
         CALL  BLKMOV
         ( SRCBLK  := "DB919_ShotResultMach".ShotResult_Ma[1],
           RET_VAL := #"Return",
           DSTBLK  := "DB919_ShotResultMach".ShotResult_Ma[0]
         );

   // Verbrauchszähler erhöhen
         CALL  "PartCounter";
         SET;
         =     "DB_Zaehler_Anzeige".Read;

         A     "DB123_MH_IO_Signals".MH[1].IN.MH_Auto_Mode;
         S     "M_NewShotDataToMC";  // For traceability
   //-
         A     "BufferShotResultM1";
         S     "DB919_ShotResultMach".ShotResult_Ma[0].General.SendData;

   m1:   NOP   0;


         AN    "DB919_ShotResultMach".ShotResult_Ma[0].General.SendData;
         R     "BufferShotResultM1";
END_REGION

REGION Network 4: PartCounter
         A     "DB_Zaehler_Anzeige".Schichtwechsel;
         JCN   Migra_CC_0;
         CALL  "PartCounterCopy";
   Migra_CC_0:SET;
         CALL  "PartCounterView";
END_REGION
END_FUNCTION_BLOCK

FUNCTION_BLOCK "FB930_FoamingData"   // FB930, STL
TITLE = Tool-Allocation -> Read tooldata and recipedata
{ S7_Optimized_Access := 'FALSE' }
AUTHOR : KT242
VERSION : 0.1
BEGIN

REGION Network 2
         CALL  "GetToolShotValues", "GetToolShotValues_DB"
         ( IN_ResetFaults    := "DB009_Faults".Faults_Reset_FKT_M1,
           IN_MachineNo      := 1,
           IN_EnableTool     := 1,
           IO_Faults         := "DB829_Error_Machine".PouringCycle[1],
           IO_FaultLevel_1   := "DB009_Faults".Faults_FKT_Grp_1_M1,
           IO_FaultLevel_2   := "DB009_Faults".Faults_FKT_Grp_2_M1,
           IO_FaultLevel_3   := "DB009_Faults".Faults_FKT_Grp_3_M1,
           IO_NewFault       := "DB009_Faults".Faultschanging_M1,
           IO_FaultAtStation := ,
           IO_PartShotNoNew  :=
         );
   //-----
END_REGION
END_FUNCTION_BLOCK

FUNCTION_BLOCK "FB1025_Service"   // FB1025, STL
{ S7_Optimized_Access := 'FALSE' }
VERSION : 0.1
   VAR_TEMP
      Inputbyte : Byte;
      Error : Word;
   END_VAR
BEGIN

REGION Network 1: Read input byte
         L     "DB1025_Service".Set.Inputbyte;
         SLW   3;
         LAR1;

         L     IB [ AR1 , P#0.0 ];
         T     "DB1025_Service".State.Inputbyte;
END_REGION

REGION Network 2: Read output byte
         L     "DB1025_Service".Set.Outputbyte;
         SLW   3;
         LAR1;

         L     QB [ AR1 , P#0.0 ];
         T     "DB1025_Service".State.Outputbyte;
END_REGION
END_FUNCTION_BLOCK

FUNCTION_BLOCK "FB1900_IF_Robots"   // FB1900, STL
TITLE = Interface Robots
{ S7_Optimized_Access := 'FALSE' }
VERSION : 0.1
   VAR_TEMP
      Auto : Bool;
      Start_cyle : Bool;
      Auto_Stop_quitt : Bool;
      Shotrelease : Bool;
      Freigabe_Eintrag_von_PUC : Bool;
      Start_Zyklus_Roboter : Bool;
      Temp_CleaningRequest : Bool;
      Temp_EnableDoorOpen : Bool;
      Automatik_Stop_ist_Quitt : Bool;
      Temp_StartCycle : Bool;
      Temp_EnableMCatPos1 : Bool;
      Temp_TestShoActiv : Bool;
      Temp_ArPos1or2 : Bool;
      Temp_FlagStartButton : Bool;
   END_VAR
BEGIN

REGION Network 1: Saftey Door 1
         ON    "DB619_State_MPart".Operationmode[1].Auto;
         ON    "DB123_MH_IO_Signals".MH[1].IN.MH_Auto_Mode;
         =     #Temp_EnableDoorOpen;
   //-----
         CALL  "FC1033_SafetyDevice"
         ( IN_With_Safety_door := true,
           IN_EnableDoorOpen   := #Temp_EnableDoorOpen,
           IN_SelectDoorOpen   := "S_SelectDoor_Robot_01",
           IN_AS_Door          := "AS_Door_Robot_01",
           IN_QuitDoorOpen     := "S_QuittDoor_Robot_01",
           IN_OMLampTest       := "DB619_State_MPart".Operationmode[1].Lamptest,
           IN_Delay_QuitDoor   := "TM_Delay_Safetydoor_1",
           OUT_V_DoorOpen      := "V_OpenDoor_Robot_01",
           OUT_H_DoorOpen      := "H_ReleaseDoor_Robot_01",
           StatusSafetyDevice  := "DB1031_AddStatus".SaftyDevice[1]
         );
   //-----
END_REGION

REGION Network 2: Saftey Door 2
         ON    "DB619_State_MPart".Operationmode[1].Auto;
         ON    "DB123_MH_IO_Signals".MH[1].IN.MH_Auto_Mode;
         =     #Temp_EnableDoorOpen;
   //-----
         CALL  "FC1033_SafetyDevice"
         ( IN_With_Safety_door := true,
           IN_EnableDoorOpen   := #Temp_EnableDoorOpen,
           IN_SelectDoorOpen   := "S_SelectDoor_TestShot_01",
           IN_AS_Door          := "AS_Door_TestShot_01",
           IN_QuitDoorOpen     := "S_QuittDoor_TestShot_01",
           IN_OMLampTest       := "DB619_State_MPart".Operationmode[1].Lamptest,
           IN_Delay_QuitDoor   := "TM_Delay_Safetydoor_2",
           OUT_V_DoorOpen      := "V_OpenDoor_TestShot_01",
           OUT_H_DoorOpen      := "H_ReleaseDoor_TestShot_01",
           StatusSafetyDevice  := "DB1031_AddStatus".SaftyDevice[2]
         );
   //-----
END_REGION

REGION Network 3: General release
         A     "AS";
         A     "DB619_State_MPart".Operationmode[1].Controllvoltage;
         A     "DB619_State_MPart".Operationmode[1].Auto;
         A     "DB123_MH_IO_Signals".MH[1].IN.MH_Auto_Mode;
         =     #Auto;
   //
         A     "AS";
         A     "DB619_State_MPart".Operationmode[1].Controllvoltage;
         =     #Auto_Stop_quitt;
   //
         AN    "AS";
         A     "DB619_State_MPart".Operationmode[1].Controllvoltage;
         A     "DB619_State_MPart".Operationmode[1].Auto;
         A     "DB123_MH_IO_Signals".MH[1].IN.MH_Auto_Mode;
         =     "DB1010_TT_Fault".AS.AS_Activ;
   //
         A     "DB619_State_MPart".Cycle[1].Release;
         =     #Shotrelease;

   // Cleaning after shot
   //-----
         A     "DB614_MH_State".MH_CleaningPiston[1].CleanAfterShotSelected;
         S     "DB1900_IF_Robots".State_Robots[1].CleaningMHRequested;
   //-
         A(;
         L     "DB1900_IF_Robots".Switch_Robots[1].StateCleaning;
         L     1;
         ==I;
         );
         R     "DB1900_IF_Robots".State_Robots[1].CleaningMHRequested;
   //-
         A     "DB1900_IF_Robots".State_Robots[1].CleaningMHRequested;
         =     #Temp_CleaningRequest;
   //-----
         CALL  "FC5901_generalFunction"
         ( StartCycle     := #Temp_StartCycle,
           EnableMCatPos1 := #Temp_EnableMCatPos1,
           TestShotActiv  := "DB1900_IF_Robots".State_Robots[1].TestShotRunning,
           AtPos1or2      := "DB1900_IF_Robots".State_Robots[1].AtPos1or2  // #Temp_ArPos1or2
         );
   //
         A     "DB1900_IF_Robots".State_Robots[1].AtPos1or2;
         =     #Temp_ArPos1or2;
END_REGION

REGION Network 4: ProgNo send to robot KUKA
         L     "DB110_Interf_Program_M1".Signals_ExPlant[1].PrgNo;
         T     "DB1900_IF_Robots".State_Kuka[1].A_SPS_PGNO;
END_REGION

REGION Network 5: Robot interface KUKA
         AN    "DB1901_Config_Robots".Config_Robots[1].Type_Kuka;
         JC    Rob_ABB;
   //------
   // Start Cycle
   //
         A     "DB110_Interf_Program_M1".Signals_ExPlant[1].cycle_run;
         FP    "FHM_PU_cycle_running";
         S     "Flag_PU_cycle_running";

         ON    "DB619_State_MPart".Cycle[1].running;
         O     "DB1900_IF_Robots".State_Kuka[1].Input_From_Robot.E_KRC_MH_OPEN;
         O     "DB1900_IF_Robots".State_Kuka[1].Input_From_Robot.E_KRC_FLT_WaitTime;
         R     "Flag_PU_cycle_running";

         A(;
         L     "DB1900_IF_Robots".State_Kuka[1].A_SPS_PGNO;
         L     0;
         >I;
         );
         A     "DB1900_IF_Robots".State_Kuka[1].Input_From_Robot.E_KRC_PGNO_REQ;
         A     "DB1900_IF_Robots".State_Kuka[1].Input_From_Robot.E_KRC_PERI_RDY;
         A     "DB1900_IF_Robots".State_Kuka[1].Input_From_Robot.E_KRC_ALARM_STOP;
         A     "DB1900_IF_Robots".State_Kuka[1].Input_From_Robot.E_KRC_USER_SAF;
         A     "DB1900_IF_Robots".State_Kuka[1].Input_From_Robot.E_KRC_AUT_EXTERN;
         A     "DB1900_IF_Robots".State_Kuka[1].Input_From_Robot.E_KRC_IN_HOME;
         A     "Flag_PU_cycle_running";
         =     #Start_cyle;


         CALL  "FC1900_IF_Kuka_KRC4"
         ( IN_PW_INOUT           := 700,
           IN_Acknowledge_Fault  := "DB009_Faults".Faults_Reset_FKT_M1,
           IN_Auto_Stop_quitt    := #Auto_Stop_quitt,
           IN_Motorprotection    := "F_Robot_01",
           IN_MH_Automatic       := #Auto,
           IN_OM_service         := "DB614_MH_State".MH_Status[1].Switch_Service_ON_OFF,
           IN_Cycle_running      := "DB619_State_MPart".Cycle[1].running,
           IN_Start_cycle        := #Start_cyle,
           IN_Release_move_MC    := TRUE,
           IN_Shotrelease        := #Shotrelease,  //"DB619_State_MPart".Cycle[1].Shotrelease
           IN_Shotend            := "DB110_Interf_Program_M1".Bits.PulseShotEnd,
           IN_FLT_Group_1        := "DB009_Faults".Fault_State_Grp_1_M1,
           IN_PGNO_MainPos       := 250,
           IN_PGNO_Cleaning      := 251,
           IN_Timer_Auto_on      := "TM_1_Robot_1",
           IN_Timer_Fault_quitt  := "TM_2_Robot_1",
           IN_Timer_Auto_On_Off  := "TM_3_Robot_1",
           IN_Timer_Delay_Start  := "TM_4_Robot_1",
           IN_Timer_PGNO_Valid   := "TM_5_Robot_1",
           IN_Timer_Imp_ExtStart := "TM_6_Robot_1",
           AB_KUKA_PGNO          := "DB1900_IF_Robots".State_Kuka[1].Output_To_Robot.A_SPS_PGNO,
           IO_Button_MainPos     := "DB1900_IF_Robots".Switch_Robots[1].SwitchMaintPosON_OFF,
           IO_Button_Cleaning    := "DB1900_IF_Robots".Switch_Robots[1].SwitchCleaningON_OFF,
           IO_State_MainPos      := "DB1900_IF_Robots".Switch_Robots[1].StateMaintPos,
           IO_State_Cleaning     := "DB1900_IF_Robots".Switch_Robots[1].StateCleaning,
           IO_Status             := "DB1900_IF_Robots".State_Kuka[1],
           IO_NewFault           := "DB009_Faults".Faultschanging_M1,
           IO_FaultLevel_3       := "DB009_Faults".Faults_FKT_Grp_3_M1
         );

   Rob_ABB:NOP   0;
END_REGION

REGION Network 6: Robot interface ABB
         AN    "DB1901_Config_Robots".Config_Robots[1].Type_ABB;
         JC    Rob_Fanuc;
   //-----
         A     "DB1900_IF_Robots".State_ABB[1].doShotDigOut_open_MH;
         A     "DB614_MH_State".MH_Status[1].OpenMHEnableExtern;
         =     "DB614_MH_State".MH_Status[1].OpenMHEnableExtern;
   //-----
   //-
         A     "DB619_State_MPart".Operationmode[1].Controllvoltage;
         =     "DB1900_IF_Robots".State_Robots[1].EmergencyStopReady;
   //-
         A     #Auto_Stop_quitt;
         =     "DB1900_IF_Robots".State_Robots[1].AutomatcStopReady;
   //-
         A     "DB619_State_MPart".Operationmode[1].Auto;
         =     "DB1900_IF_Robots".State_Robots[1].MaschineAuto;
   //-
         A     "DB123_MH_IO_Signals".MH[1].IN.MH_Auto_Mode;
         =     "DB1900_IF_Robots".State_Robots[1].MixingheadAuto;
   //-
   // Status auch in FC irgendwann!

         A     "DB1900_IF_Robots".State_ABB[1].Output.doIRBInHome;
         =     "DB1900_IF_Robots".State_Robots[1].Rob_in_Home;

         A     "DB1900_IF_Robots".State_ABB[1].Output.doIRBinAuto;
         =     "DB1900_IF_Robots".State_Robots[1].Rob_in_Automatic;

         A     "DB1900_IF_Robots".State_ABB[1].Output.doCycleStarted;
         =     "DB1900_IF_Robots".State_Robots[1].Rob_in_Cycle;

         A     "DB1900_IF_Robots".State_ABB[1].Output.doIRBinAuto;
         A     "DB1900_IF_Robots".State_ABB[1].Output.doIRBInHome;
         A     "DB1900_IF_Robots".State_ABB[1].Output.doCycleEnd;
         A(;
         L     "DB1900_IF_Robots".State_ABB[1].Stepnumber;
         L     0;
         ==I;
         );
         =     "DB1900_IF_Robots".State_Robots[1].ReadyForStartCycle;

         L     "DB1900_IF_Robots".State_ABB[1].Stepnumber;
         T     "DB1900_IF_Robots".State_Robots[1].StepNo;

         L     "DB1900_IF_Robots".State_ABB[1].Output.GOError;
         T     "DB1900_IF_Robots".State_Robots[1].FaultNo;
   ///----------
   // Not- Aus und Automatik Stop wurden quittiert:
   ///----------
         AN    "DB1900_IF_Robots".State_ABB[1].Output.doSysError;
         AN    "DB1900_IF_Robots".State_ABB[1].Output.doEmStop_Akt;
         AN    "DB1900_IF_Robots".State_ABB[1].Input.diQuickStop;
         AN    "DB1900_IF_Robots".State_ABB[1].Output.doSafeZoneActiv;
         A     #Auto_Stop_quitt;
         A     "DB123_MH_IO_Signals".MH[1].IN.MH_Auto_Mode;
         =     #Automatik_Stop_ist_Quitt;
   ///----------
   // Datenaustausch mit dem Roboter starten:
   ///----------
         A     #Temp_StartCycle;
         A     #Automatik_Stop_ist_Quitt;
         A     "DB1900_IF_Robots".State_ABB[1].Output.doIRBInHome;
         A     "DB1900_IF_Robots".State_ABB[1].Output.doIRBinAuto;
         A     "DB1900_IF_Robots".State_ABB[1].Output.doCycleOn;
         AN    "DB1900_IF_Robots".State_ABB[1].Output.doSysError;
         AN    "DB619_State_MPart".Operationmode[1].Test;
         =     #Start_Zyklus_Roboter;
   ///----------
   // Bewegungefreigabe zum Verfahren in die Formträger
   ///----------
         A     #Temp_EnableMCatPos1;
         A     "DB123_MH_IO_Signals".MH[1].IN.MH_Auto_Mode;
         AN    "DB619_State_MPart".Operationmode[1].Test;
         A     "DB619_State_MPart".Cycle[1].Shotrelease;
   //U     "DB005_RS<->Extern".MC_Interface[1].FromMC.EnableFoaming
         =     "DB1900_IF_Robots".State_ABB[1].Input.diStartMoveMC;
   //--------------------------------------------------------------------
   // Das öffnen des Mischkopfes kann von dem Roboter angesteuert werden:
   // Roboter wartet in Vorposition bis das Signal kommt.
         A     #Temp_EnableMCatPos1;
         A     "DB619_State_MPart".Cycle[1].Shotrelease;
         =     #Freigabe_Eintrag_von_PUC;
   ///----------
   // Roboter zur Maintenanceposition und zurück zur Homeposition
   ///----------
         A     "DB1900_IF_Robots".Switch_Robots[1].SwitchMaintPosON_OFF;
         A     "DB123_MH_IO_Signals".MH[1].IN.MH_Auto_Mode;
         AN    #Temp_ArPos1or2;
         A     #Automatik_Stop_ist_Quitt;  // NotHalt ???
         A     "DB1900_IF_Robots".State_ABB[1].Output.doIRBInHome;
         A     "DB1900_IF_Robots".State_ABB[1].Output.doCycleEnd;
         AN    "DB1900_IF_Robots".State_ABB[1].Output.doCycleStarted;
         S     "DB1900_IF_Robots".State_ABB[1].Input.diHomeToMaintP;
   ///----------
         O     "DB1900_IF_Robots".State_ABB[1].Output.doIRBInMaintP;
         ON    "DB1900_IF_Robots".State_ABB[1].Output.doIRBinAuto;
         ON    "DB1900_IF_Robots".State_ABB[1].Output.doCycleOn;
         R     "DB1900_IF_Robots".State_ABB[1].Input.diHomeToMaintP;
   ///----------
         AN    "DB1900_IF_Robots".Switch_Robots[1].SwitchMaintPosON_OFF;
         A     "DB123_MH_IO_Signals".MH[1].IN.MH_Auto_Mode;
         A     #Automatik_Stop_ist_Quitt;
         A     "DB1900_IF_Robots".State_ABB[1].Output.doIRBInMaintP;
         A     "DB1900_IF_Robots".State_ABB[1].Output.doCycleEnd;
         AN    "DB1900_IF_Robots".State_ABB[1].Output.doCycleStarted;
         S     "DB1900_IF_Robots".State_ABB[1].Input.diMaintToHomeP;
   ///----------
         O     "DB1900_IF_Robots".State_ABB[1].Output.doIRBInHome;
         ON    "DB1900_IF_Robots".State_ABB[1].Output.doIRBinAuto;
         ON    "DB1900_IF_Robots".State_ABB[1].Output.doCycleOn;
         R     "DB1900_IF_Robots".State_ABB[1].Input.diMaintToHomeP;
   //-----
         L     1;  // Green
         A     "DB1900_IF_Robots".State_ABB[1].Output.doIRBInMaintP;
         JC    StateMaintPos;
         L     3;  // Yellow
         O     "DB1900_IF_Robots".Switch_Robots[1].SwitchMaintPosON_OFF;
         O     "DB1900_IF_Robots".State_ABB[1].Input.diMaintToHomeP;
         JC    StateMaintPos;
         L     0;  // OFF
   StateMaintPos:NOP   0;
         T     "DB1900_IF_Robots".Switch_Robots[1].StateMaintPos;

   ///----------
   // Roboter zur 2. Maintenanceposition und zurück zur Homeposition
   ///----------
         A     "DB1900_IF_Robots".Switch_Robots[1].SwitchMaintPos_2ON_OFF;
         A     "DB123_MH_IO_Signals".MH[1].IN.MH_Auto_Mode;
         AN    #Temp_ArPos1or2;
         A     #Automatik_Stop_ist_Quitt;  // NotHalt ???
         A     "DB1900_IF_Robots".State_ABB[1].Output.doIRBInHome;
         A     "DB1900_IF_Robots".State_ABB[1].Output.doCycleEnd;
         AN    "DB1900_IF_Robots".State_ABB[1].Output.doCycleStarted;
         S     "DB1900_IF_Robots".State_ABB[1].Input.diHomeToMaint2;
   ///----------
         O     "DB1900_IF_Robots".State_ABB[1].Output.doIRBInMaintP2;
         ON    "DB1900_IF_Robots".State_ABB[1].Output.doIRBinAuto;
         ON    "DB1900_IF_Robots".State_ABB[1].Output.doCycleOn;
         R     "DB1900_IF_Robots".State_ABB[1].Input.diHomeToMaint2;
   ///----------
         AN    "DB1900_IF_Robots".Switch_Robots[1].SwitchMaintPos_2ON_OFF;
         A     "DB123_MH_IO_Signals".MH[1].IN.MH_Auto_Mode;
         A     #Automatik_Stop_ist_Quitt;
         A     "DB1900_IF_Robots".State_ABB[1].Output.doIRBInMaintP2;
         A     "DB1900_IF_Robots".State_ABB[1].Output.doCycleEnd;
         AN    "DB1900_IF_Robots".State_ABB[1].Output.doCycleStarted;
         S     "DB1900_IF_Robots".State_ABB[1].Input.diMaintToHome2;
   ///----------
         O     "DB1900_IF_Robots".State_ABB[1].Output.doIRBInHome;
         ON    "DB1900_IF_Robots".State_ABB[1].Output.doIRBinAuto;
         ON    "DB1900_IF_Robots".State_ABB[1].Output.doCycleOn;
         R     "DB1900_IF_Robots".State_ABB[1].Input.diMaintToHome2;
   //-----

         L     1;  // Green
         A     "DB1900_IF_Robots".State_ABB[1].Output.doIRBInMaintP2;
         JC    StateMaintPos2;
         L     3;  // Yellow
         O     "DB1900_IF_Robots".Switch_Robots[1].SwitchMaintPos_2ON_OFF;
         O     "DB1900_IF_Robots".State_ABB[1].Input.diMaintToHome2;
         JC    StateMaintPos2;
         L     0;  // OFF
   StateMaintPos2:NOP   0;
         T     "DB1900_IF_Robots".Switch_Robots[1].StateMaintPos_2;

   //-----
   // Robot to mixinghead cleaning
   //-----
         A(;
         A     "DB1900_IF_Robots".Switch_Robots[1].SwitchBrushON_OFF;
         AN    #Temp_ArPos1or2;
         A     "DB1900_IF_Robots".State_ABB[1].Output.doIRBInHome;
         A     "DB1900_IF_Robots".State_ABB[1].Output.doCycleEnd;
         AN    "DB1900_IF_Robots".State_ABB[1].Output.doCycleStarted;
         O;
         A     "DB619_State_MPart".Cycle[1].ShotRuns;
         A     "DB614_MH_State".MH_CleaningPiston[1].CleanAfterShotSelected;
         );
         A     #Automatik_Stop_ist_Quitt;
         S     "DB1900_IF_Robots".State_ABB[1].Input.diStartBrushMH;
         S     "DB1900_IF_Robots".State_ABB[1].CleaningSelected;
   //-----
         O     "DB1900_IF_Robots".State_ABB[1].Output.doCleanBrushOn;
         ON    "DB1900_IF_Robots".State_ABB[1].Output.doIRBinAuto;
         ON    "DB1900_IF_Robots".State_ABB[1].Output.doCycleOn;
         R     "DB1900_IF_Robots".State_ABB[1].Input.diStartBrushMH;
   //-----
         A     "DB1900_IF_Robots".State_ABB[1].Output.doCleanBrushOn;
         FN    "DB1900_IF_Robots".State_ABB[1].FHM_CleaningActiv;
         =     "DB1900_IF_Robots".State_ABB[1].CleaningActiv;
   //-----
         A     "DB1900_IF_Robots".State_ABB[1].CleaningActiv;
         R     "DB1900_IF_Robots".State_ABB[1].CleaningSelected;
         R     "DB1900_IF_Robots".Switch_Robots[1].SwitchBrushON_OFF;
   //-----
   // Ansteuerung des Reinigungskolben vom Roboter aus
         A     "DB1900_IF_Robots".State_ABB[1].Output.doCleanBrushOn;
         =     "DB1900_IF_Robots".State_Robots[1].CleaningMHOn;
   //-----
         L     1;  // Green
         A     "DB1900_IF_Robots".State_ABB[1].Output.doCleanBrushOn;
         JC    StateCleaningMH;
         L     3;  // Yellow
         O     "DB1900_IF_Robots".Switch_Robots[1].SwitchBrushON_OFF;
         O     "DB1900_IF_Robots".State_ABB[1].CleaningSelected;
         JC    StateCleaningMH;
         L     0;  // OFF
   StateCleaningMH:NOP   0;
         T     "DB1900_IF_Robots".Switch_Robots[1].StateBrush;

   //-----
   // Robot to Synchronize EPS
   //-----
         A     "DB1900_IF_Robots".State_ABB[1].Output.doSafetyPreWarn;
         A     "DB1900_IF_Robots".State_ABB[1].Output.doIRBinAuto;
         A     "DB123_MH_IO_Signals".MH[1].IN.MH_Auto_Mode;
         O     "DB1900_IF_Robots".Switch_Robots[1].SwitchSyncON_OFF;
         FP    "DB1900_IF_Robots".State_ABB[1].FHM_SyncEPS;
         S     "DB1900_IF_Robots".State_ABB[1].Start_Synchronization;
   //-----
         A     "DB1900_IF_Robots".State_ABB[1].Start_Synchronization;
         A     #Automatik_Stop_ist_Quitt;
         AN    "DB619_State_MPart".Cycle[1].running;
         AN    #Temp_ArPos1or2;
         A     "DB1900_IF_Robots".State_ABB[1].Output.doIRBInHome;
         A     "DB1900_IF_Robots".State_ABB[1].Output.doIRBinAuto;
         A     "DB1900_IF_Robots".State_ABB[1].Output.doCycleEnd;
         AN    "DB1900_IF_Robots".State_ABB[1].Output.doCycleStarted;
         =     "DB1900_IF_Robots".State_ABB[1].Input.diStartSyncSafety;
   //-----
         O     "DB1900_IF_Robots".State_ABB[1].Output.doSafetySyncSwitch;
         O     "DB1900_IF_Robots".State_ABB[1].Output.doSafetyControlPos;
         O     "Flag_Erster_SPS_Zyklus";
         R     "DB1900_IF_Robots".State_ABB[1].Input.diStartSyncSafety;
         R     "DB1900_IF_Robots".State_ABB[1].Start_Synchronization;
         R     "DB1900_IF_Robots".Switch_Robots[1].SwitchSyncON_OFF;
   //-----
         L     1;  // Green
         A     "DB1900_IF_Robots".State_ABB[1].Output.doSafetySynchronized;
         AN    "DB1900_IF_Robots".State_ABB[1].Start_Synchronization;
         JC    StateSync;
         L     3;
         A     "DB1900_IF_Robots".State_ABB[1].Start_Synchronization;
         JC    StateSync;
         L     2;  // Red
   StateSync:NOP   0;
         T     "DB1900_IF_Robots".Switch_Robots[1].StateSync;
   //-----
   //    Störung:
   //-----
         A     "DB009_Faults".Faults_Reset_FKT_M1;
         R     "DB1900_IF_Robots".Faults_Robots[1].FLT_SyncPosition;
   //---
         AN    "DB1900_IF_Robots".State_ABB[1].Output.doSafetySyncSwitch;
         A     "DB1900_IF_Robots".State_ABB[1].Output.doSafetyControlPos;
         L     S5T#1S;
         SD    "TM_Verz_Sync_1";
         A     "TM_Verz_Sync_1";
         AN    "DB1900_IF_Robots".Faults_Robots[1].FLT_SyncPosition;
         S     "DB1900_IF_Robots".Faults_Robots[1].FLT_SyncPosition;
         S     "DB009_Faults".Faultschanging_M1;
         A     "DB1900_IF_Robots".Faults_Robots[1].FLT_SyncPosition;
         S     "DB009_Faults".Faults_FKT_Grp_1_M1;
   //------------------------------------------------------------------
         AN    "DB1900_IF_Robots".State_ABB[1].Output.doSafeZoneActiv;
         =     "Tag_3";
         =     "Tag_4";

         CLR;
         =     "DB1900_IF_Robots".State_ABB[1].Input.diQuickStop;

         SET;
         =     "DB1900_IF_Robots".State_ABB[1].Input.diRobinSavepos;
   //-----
   //Daten Roboterabhängig kopieren
         L     "DB110_Interf_Program_M1".Robot_01.Robot_ProgNo_Mould_1;
         T     "DB1900_IF_Robots".State_ABB[1].Robot_ProgNo_Mould_1;
         L     "DB110_Interf_Program_M1".Robot_01.Robot_ProgNo_Mould_2;
         T     "DB1900_IF_Robots".State_ABB[1].Robot_ProgNo_Mould_2;
         L     "DB110_Interf_Program_M1".Robot_01.Robot_ProgNo_Mould_3;
         T     "DB1900_IF_Robots".State_ABB[1].Robot_ProgNo_Mould_3;

         L     "DB110_Interf_Program_M1".Robot_01.MC_Place_Number;
         T     "DB1900_IF_Robots".State_ABB[1].MC_Place_Number;
         T     "DB1900_IF_Robots".State_Fanuc[1].MCPlaceNumber;
   //-----
         CALL  "FC1910_IF_ABB"
         ( IN_PW_Ein_Ausgaenge      := 600,
           IN_Reset_fault_Fkt       := "DB009_Faults".Faults_Reset_FKT_M1,
           IN_Steuerspannung        := "DB619_State_MPart".Operationmode[1].Controllvoltage,
           IN_Zyklus_Laeuft         := "DB619_State_MPart".Cycle[1].running,
           IN_Zyklus_KLZ1_Laeuft    := "DB619_State_MPart".Cycle[1].PressurizeTimeRuns,
           IN_Zyklus_KLZ3_Laeuft    := "DB619_State_MPart".Cycle[1].StandByTimeRuns,
           IN_Zyklus_Schuss_laeuft  := "DB619_State_MPart".Cycle[1].ShotRuns,
           IN_Imp_Schussende        := "DB619_State_MPart".Cycle[1].PulsShotend,
           IN_Imp_Prog_Letzter_TS   := FALSE,
           IN_Betriebsart_Automatik := "DB619_State_MPart".Operationmode[1].Auto,
           IN_MK_Automatik          := "DB123_MH_IO_Signals".MH[1].IN.MH_Auto_Mode,
           IN_Anf_Flucht            := FALSE,
           IN_Auto_Stop_quittiert   := #Automatik_Stop_ist_Quitt,
           IN_Zyklus_Freigabe       := "DB619_State_MPart".Cycle[1].Release,
           IN_Zyklus_Max_Wartezeit  := "DB619_State_MPart".Cycle[1].FLT_MaxWaittime,
           IN_Start_Prog_Imp        := #Start_Zyklus_Roboter,
           IN_FRG_Datatransfer      := TRUE,
           IN_FRG_von_PU            := #Freigabe_Eintrag_von_PUC,
           IN_Anwahl_Mit_Shotware   := FALSE,
           IN_Anwahl_Mit_Tracking   := FALSE,
           IN_Timer_Auto_ein_Track  := "TM_1_Robot_1",
           IN_Timer_Auto_ein        := "TM_2_Robot_1",
           IN_Timer_Verz_Handanwahl := "TM_3_Robot_1",
           IN_Timer_Auto_aus        := "TM_4_Robot_1",
           IN_Timer_Fluchtprog      := "TM_5_Robot_1",
           IN_Timer_Start_Verz      := "TM_6_Robot_1",
           IN_Timer_Start_Main_Verz := "TM_7_Robot_1",
           IN_Schusszeit            := w#16#0,  //"DB111_ShotvaluesRobot_M1"
           IO_Status                := "DB1900_IF_Robots".State_ABB[1],
           IO_Fault                 := "DB1900_IF_Robots".Faults_Robots[1],
           IO_NewFault              := "DB009_Faults".Faultschanging_M1,
           IO_FaultLevel_1          := "DB009_Faults".Faults_FKT_Grp_1_M1,
           IO_FaultLevel_2          := "DB009_Faults".Faults_FKT_Grp_2_M1,
           IO_FaultLevel_3          := "DB009_Faults".Faults_FKT_Grp_3_M1
         );

   // Fault handling
   //------------------------------------------------------------------
   //      U     "DB009_Faults".Faults_Reset_FKT_M1
   //      R     "DB1900_IF_Robots".Faults_Robots[1].FLT_Fuse
   //      R     "DB825_Error_Interface".Roboter[1].FLT_Stepnumber_not_zero

   //--      UN    "F_Supply_Roboter"
   //--      UN    "DB1900_IF_Robots".Faults_Robots[1].FLT_Fuse
   //--      S    "DB1900_IF_Robots".Faults_Robots[1].FLT_Fuse
   //--      S     "DB009_Faults".Faultschanging_M1
   //---
   //      U     "DB1900_IF_Robots".State_ABB[1].Output.doIRBinAuto
   //      U     "DB1900_IF_Robots".State_ABB[1].Output.doIRBInHome
   //      U     "DB1900_IF_Robots".State_ABB[1].Output.doCycleEnd
   //      U(
   //      L     "DB1900_IF_Robots".State_ABB[1].Stepnumber
   //      L     0
   //      <>I
   //      )
   //      L     S5T#3S
   //--      SE    "TM_F_Schrittnummer_Rob01"

   //--      U     "TM_F_Schrittnummer_Rob01"
   //      UN    "DB825_Error_Interface".Roboter[1].FLT_Stepnumber_not_zero
   //      S     "DB825_Error_Interface".Roboter[1].FLT_Stepnumber_not_zero
   //      S     "DB009_Faults".Faultschanging_M1

   //      O     "DB1900_IF_Robots".Faults_Robots[1].FLT_Fuse
   //      O     "DB825_Error_Interface".Roboter[1].FLT_Stepnumber_not_zero
   //      S     "DB009_Faults".Faults_FKT_Grp_3_M1
   //_________________________________________________________________________


   //  Messages:
   //-------------------------------------------------------------------------
   //      U     #Automatik_Stop_ist_Quitt
   //      U     "DB1900_IF_Robots".State_ABB[1].Output.doIRBinAuto
   //      UN    "DB1900_IF_Robots".State_ABB[1].Output.doCycleOn
   //      UN    "DB1900_IF_Robots".State_ABB[1].Output.doSysError
   //      L     S5T#10S
   //--      SE    "TM_STG_Rob1_Prg"
   //--      U     "TM_STG_Rob1_Prg"
   //--      =     "RobNotRunning"

   //--      U     "RobNotRunning"
   //      UN    "DB825_Error_Interface".Roboter[1].RobotProgramNotRunning
   //      S     "DB825_Error_Interface".Roboter[1].RobotProgramNotRunning
   //      S     "DB009_Faults".NewMessage_M1

   //--      UN    "RobNotRunning"
   //      R     "DB825_Error_Interface".Roboter[1].RobotProgramNotRunning
   //      S     "DB009_Faults".GoneMessage_M1


         A     "DB619_State_MPart".Operationmode[1].Controllvoltage;
         A     "DB619_State_MPart".Operationmode[1].Auto;
         A     "DB123_MH_IO_Signals".MH[1].IN.MH_Auto_Mode;
         AN    "DB1900_IF_Robots".State_ABB[1].Output.doIRBinAuto;
         =     "DB1900_IF_Robots".Faults_Robots[1].MSG_Rob_not_in_automatic;
   //_________________________________________________________________________
   //
   Rob_Fanuc:NOP   0;
END_REGION

REGION Network 7: Robot interface Fanuc
         AN    "DB1901_Config_Robots".Config_Robots[1].Type_Fanuc;
         JC    Rob_Motoman;

   // Datenaustausch mit dem Roboter starten:
   //
         O     "DB110_Interf_Program_M1".Status_IF[1].Start_to_Cycle;  //Start from OP-Panel or mouldcarrier
         O     "DB110_Interf_Program_M1".Status_IF[2].Start_to_Cycle;  //Start from OP-Panel or mouldcarrier
         O     "DB110_Interf_Program_M1".Status_IF[3].Start_to_Cycle;  //Start from OP-Panel or mouldcarrier
         A     "DB123_MH_IO_Signals".MH[1].IN.MH_Auto_Mode;
         A     "DB1900_IF_Robots".State_Fanuc[1].Output.do_IRB_Auto;
         A     "DB1900_IF_Robots".State_Fanuc[1].Output.SYSRDY_Robot_sys_ready;
         AN    "DB1900_IF_Robots".State_Fanuc[1].Output.Fault_Robot;
         AN    "DB619_State_MPart".Operationmode[1].Test;
         =     #Start_Zyklus_Roboter;

   ///----------
   // Bewegungsfreigabe zum Verfahren in die Formträger
   ///----------

         O     "DB110_Interf_Program_M1".Status_IF[1].IF_is_on_1_Position;
         O     "DB110_Interf_Program_M1".Status_IF[2].IF_is_on_1_Position;
         A     "DB123_MH_IO_Signals".MH[1].IN.MH_Auto_Mode;
         AN    "DB619_State_MPart".Operationmode[1].Test;
         A(;
         O     "DB1900_IF_Robots".State_Fanuc[1].Output.goFormAktBit0;
         O     "DB1900_IF_Robots".State_Fanuc[1].Output.goFormAktBit1;
         );
         =     "DB1900_IF_Robots".State_Fanuc[1].Input.diRelMoveMC;

   //-----------
   // Freigabe für die HomePos- Fahrt
   //-----------
         SET;
         =     "DB1900_IF_Robots".State_Fanuc[1].Input.diEnableHome;
   //
   //--------------------------------------------------------------------
   // Das öffnen des Mischkopfes kann von dem Roboter angesteuert werden:
   // Roboter wartet in Vorposition bis das Signal kommt.
         A(;
         O     "DB110_Interf_Program_M1".Status_IF[1].IF_is_on_1_Position;
         O     "DB110_Interf_Program_M1".Status_IF[2].IF_is_on_1_Position;
         O     "DB110_Interf_Program_M1".Status_IF[3].IF_is_on_1_Position;
         );
         A     "DB619_State_MPart".Cycle[1].Shotrelease;  //Pressure build up- or control time finished
         A     "DB619_State_MPart".Mixinghead[1].Cleaningpiston_OK;
         =     #Freigabe_Eintrag_von_PUC;

   //Daten Roboterabhängig kopieren
         L     "DB110_Interf_Program_M1".Robot_01.Robot_ProgNo_Mould_1;
         T     "DB1900_IF_Robots".State_Fanuc[1].RobotProgNoMould1;
         L     "DB110_Interf_Program_M1".Robot_01.Robot_ProgNo_Mould_2;
         T     "DB1900_IF_Robots".State_Fanuc[1].RobotProgNoMould2;
         L     "DB110_Interf_Program_M1".Robot_01.Robot_ProgNo_Mould_3;
         T     "DB1900_IF_Robots".State_Fanuc[1].RobotProgNoMould3;

         L     "DB110_Interf_Program_M1".Robot_01.MC_Place_Number;
         T     "DB1900_IF_Robots".State_Fanuc[1].MCPlaceNumber;

   // Ansteuerung des Reinigungskolben vom Roboter aus
         A     "DB1900_IF_Robots".State_Fanuc[1].Output.doCleaningPLC;
         =     "DB1900_IF_Robots".State_Robots[1].CleaningMHOn;
   //-----
         CALL  "FC1920_IF_Fanuc"
         ( IN_AdressRobIO           := 300,
           IN_ResetFaultFct         := "DB009_Faults".Faults_Reset_FKT_M1,
           IN_ControlVoltage        := "DB619_State_MPart".Operationmode[1].Controllvoltage,
           IN_FoamingCycleRunning   := "DB619_State_MPart".Cycle[1].running,
           IN_MHAutomatic           := #Auto,
           IN_RequestEscapeProg     := FALSE,
           IN_AutoStopOK            := #Auto_Stop_quitt,
           IN_FuseSupplyOK          := "F_Robot_01",
           IN_EnableFoamingCycle    := #Shotrelease,
           IN_ShotActive            := "DB619_State_MPart".Cycle[1].ShotRuns,
           IN_CycleMaxWaitingTime   := "DB619_State_MPart".Cycle[1].FLT_MaxWaittime,
           IN_StartPulseDataExchang := #Start_Zyklus_Roboter,
           IN_PulseShotEnd          := "DB110_Interf_Program_M1".Bits.PulseShotEnd,
           IN_EnableDataExchange    := TRUE,
           IN_EnableShotFromPU      := #Freigabe_Eintrag_von_PUC,
           IN_ConfigWithTracking    := "DB1901_Config_Robots".Config_Robots[1].With_Tracking,
           IN_OtherRobotOnly        := FALSE,
           IN_CleaningRequest       := #Temp_CleaningRequest,
           IN_PGNO_MainPos          := 1003,
           IN_PGNO_MainPos2         := 0,
           IN_PGNO_Cleaning         := 1000,
           IN_PGNO_Testshot         := 1005,
           IN_TimerAutoOnTrack      := "TM_1_Robot_1",
           IN_TimerAutoOn           := "TM_2_Robot_1",
           IN_TimerDelayManSelect   := "TM_3_Robot_1",
           IN_TimerAutoOFF          := "TM_4_Robot_1",
           IN_TimerEscapeProg       := "TM_5_Robot_1",
           IN_TimerStartDelay       := "TM_6_Robot_1",
           IN_TimerFaultReset       := "TM_7_Robot_1",
           IO_Button_MainPos        := "DB1900_IF_Robots".Switch_Robots[1].SwitchMaintPosON_OFF,
           IO_Button_MainPos2       := "DB1900_IF_Robots".Switch_Robots[1].SwitchMaintPos_2ON_OFF,
           IO_Button_Cleaning       := "DB1900_IF_Robots".Switch_Robots[1].SwitchCleaningON_OFF,
           IO_Button_Testshot       := "DB1900_IF_Robots".Switch_Robots[1].SwitchTestShotON_OFF,
           IO_State_MainPos         := "DB1900_IF_Robots".Switch_Robots[1].StateMaintPos,
           IO_State_MainPos2        := "DB1900_IF_Robots".Switch_Robots[1].StateMaintPos_2,
           IO_State_Cleaning        := "DB1900_IF_Robots".Switch_Robots[1].StateCleaning,
           IO_State_Testshot        := "DB1900_IF_Robots".Switch_Robots[1].StateTestShot,
           IO_Status                := "DB1900_IF_Robots".State_Fanuc[1],
           IO_NewFault              := "DB009_Faults".Faultschanging_M1,
           IO_FaultLevel_1          := "DB009_Faults".Faults_FKT_Grp_1_M1,
           IO_FaultLevel_3          := "DB009_Faults".Faults_FKT_Grp_3_M1,
           IO_Faults                := "DB1900_IF_Robots".State_Fanuc[1].Faults
         );

   Rob_Motoman:NOP   0;
END_REGION

REGION Network 8: Robot interface Motoman
         AN    "DB1901_Config_Robots".Config_Robots[1].Type_Motoman;
         JC    End;
END_REGION

REGION Network 9: End / Copy Faults to general Fault state
   // Erstmal so. Soll eigtl. direkt in die FCs
   End:  NOP   0;

         A     "DB1901_Config_Robots".Config_Robots[1].Type_ABB;
         JC    NoFunction;

         A     "DB1900_IF_Robots".State_Fanuc[1].Faults.FLT_System;
         A     "DB1901_Config_Robots".Config_Robots[1].Type_Fanuc;
         O;
         A     "DB1900_IF_Robots".State_Kuka[1].STG_System;
         A     "DB1901_Config_Robots".Config_Robots[1].Type_Kuka;
         =     "DB1900_IF_Robots".Faults_Robots[1].FLT_System;

         A     "DB1900_IF_Robots".State_Fanuc[1].Faults.FLT_Interface;
         A     "DB1901_Config_Robots".Config_Robots[1].Type_Fanuc;
         O;
         A     "DB1900_IF_Robots".State_Kuka[1].STG_Schnittstelle;
         A     "DB1901_Config_Robots".Config_Robots[1].Type_Kuka;
         =     "DB1900_IF_Robots".Faults_Robots[1].FLT_Interface;

         A     "DB1900_IF_Robots".State_Fanuc[1].Faults.FLT_RobStoppedInProd;
         A     "DB1901_Config_Robots".Config_Robots[1].Type_Fanuc;
         O;
         A     "DB1900_IF_Robots".State_Kuka[1].STG_Roboter_stoppt;
         A     "DB1901_Config_Robots".Config_Robots[1].Type_Kuka;
         =     "DB1900_IF_Robots".Faults_Robots[1].FLT_Prog_stopped;

         A     "DB1900_IF_Robots".State_Fanuc[1].Faults.FLT_Fuse_Supply;
         A     "DB1901_Config_Robots".Config_Robots[1].Type_Fanuc;
         O;
         A     "DB1900_IF_Robots".State_Kuka[1].STG_Motoschutz;
         A     "DB1901_Config_Robots".Config_Robots[1].Type_Kuka;
         =     "DB1900_IF_Robots".Faults_Robots[1].FLT_Fuse;

         A     "DB1900_IF_Robots".State_Fanuc[1].Faults.FLT_PrgNotExisting;
         A     "DB1901_Config_Robots".Config_Robots[1].Type_Fanuc;

         =     "DB1900_IF_Robots".Faults_Robots[1].FLT_Wrong_Prog_No;
         CLR;
         =     "DB1900_IF_Robots".Faults_Robots[1].FLT_Wrong_MC_No;
         CLR;
         =     "DB1900_IF_Robots".Faults_Robots[1].FLT_Wrong_Shot_time;
         A     "DB1900_IF_Robots".State_Fanuc[1].Faults.FLT_TPOnInProd;
         A     "DB1901_Config_Robots".Config_Robots[1].Type_Fanuc;

         =     "DB1900_IF_Robots".Faults_Robots[1].FLT_TP_On_in_automatic;


         A     "DB1900_IF_Robots".State_Fanuc[1].Faults.Roboter_not_in_automatic;
         A     "DB1901_Config_Robots".Config_Robots[1].Type_Fanuc;
         O;
         A     "DB1900_IF_Robots".State_Kuka[1].Anforderung_Automatik;
         A     "DB1901_Config_Robots".Config_Robots[1].Type_Kuka;

         =     "DB1900_IF_Robots".Faults_Robots[1].MSG_Rob_not_in_automatic;
         CLR;
         =     "DB1900_IF_Robots".Faults_Robots[1].MSG_Emergency_stop_Robot;


   // Status auch in FC irgendwann!


   NoFunction:NOP   0;

         A     "DB009_Faults".Faults_Reset_FKT_M1;
         R     "DB1900_IF_Robots".Faults_Robots[1].FLT_Fuse;

         AN    "F_Robot_01";
         AN    "DB1900_IF_Robots".Faults_Robots[1].FLT_Fuse;
         CLR;
         S     "DB1900_IF_Robots".Faults_Robots[1].FLT_Fuse;
         S     "DB009_Faults".Faultschanging_M1;
         S     "DB009_Faults".Faults_FKT_Grp_3_M1;

         AN    "ES_Robot_01";
         =     "DB1900_IF_Robots".Faults_Robots[1].MSG_Emergency_stop_Robot;

         A     "DB1900_IF_Robots".State_Fanuc[1].Output.doIRBInHome;
         A     "DB1901_Config_Robots".Config_Robots[1].Type_Fanuc;
         O;
         A     "DB1900_IF_Robots".State_ABB[1].Output.doIRBInHome;
         A     "DB1901_Config_Robots".Config_Robots[1].Type_ABB;

         =     "DB1900_IF_Robots".State_Robots[1].Rob_in_Home;

         A     "DB1900_IF_Robots".State_Fanuc[1].AutomaticAccepted;
         A     "DB1901_Config_Robots".Config_Robots[1].Type_Fanuc;
         O;
         A     "DB1900_IF_Robots".State_ABB[1].Auto_accepted;
         A     "DB1901_Config_Robots".Config_Robots[1].Type_ABB;

         =     "DB1900_IF_Robots".State_Robots[1].Rob_in_Automatic;

         A     "DB1900_IF_Robots".State_Fanuc[1].StartFoamingCycle;
         A     "DB1901_Config_Robots".Config_Robots[1].Type_Fanuc;
         O;
         A     "DB1900_IF_Robots".State_ABB[1].Output.doCycleStarted;
         A     "DB1901_Config_Robots".Config_Robots[1].Type_ABB;

         =     "DB1900_IF_Robots".State_Robots[1].Rob_in_Cycle;

         L     "DB110_Interf_Program_M1".Robot_01.Robot_ProgNo_Mould_1;
         T     "DB1900_IF_Robots".State_Robots[1].Rob_Prog_No;

         L     "DB110_Interf_Program_M1".Robot_01.MC_Place_Number;
         T     "DB1900_IF_Robots".State_Robots[1].Rob_MC_No;
END_REGION

REGION Network 10: Delete faults if no robot is selected
         AN    "DB1901_Config_Robots".Config_Robots[1].Type_Kuka;
         AN    "DB1901_Config_Robots".Config_Robots[1].Type_ABB;
         AN    "DB1901_Config_Robots".Config_Robots[1].Type_Fanuc;
         AN    "DB1901_Config_Robots".Config_Robots[1].Type_Motoman;
         R     "DB1900_IF_Robots".Faults_Robots[1].FLT_System;
         R     "DB1900_IF_Robots".Faults_Robots[1].FLT_Interface;
         R     "DB1900_IF_Robots".Faults_Robots[1].FLT_Prog_stopped;
   //      R     "DB1900_IF_Robots".Faults_Robots[1].FLT_Fuse
         R     "DB1900_IF_Robots".Faults_Robots[1].FLT_Wrong_Prog_No;
         R     "DB1900_IF_Robots".Faults_Robots[1].FLT_Wrong_MC_No;
         R     "DB1900_IF_Robots".Faults_Robots[1].FLT_TP_On_in_automatic;
         R     "DB1900_IF_Robots".Faults_Robots[1].MSG_Rob_not_in_automatic;
         R     "DB1900_IF_Robots".Faults_Robots[1].MSG_Emergency_stop_Robot;
END_REGION
END_FUNCTION_BLOCK

FUNCTION_BLOCK "GetToolShotValues"   // FB1930, SCL
TITLE = Get shotvalues from selected tool
{ S7_Optimized_Access := 'FALSE' }
VERSION : 0.1
   VAR_INPUT
      IN_ResetFaults : Bool;
      IN_MachineNo : Int;
      IN_EnableTool : Bool;
   END_VAR
   VAR_IN_OUT
      IO_Faults : "UDT1819_FLT_PouringCycle";
      IO_FaultLevel_1 : Bool;   // Fault message of level 1 is active and was not acknowledged
      IO_FaultLevel_2 : Bool;   // Fault message of level 2 is active and was not acknowledged
      IO_FaultLevel_3 : Bool;   // Fault message of level 3 is active and was not acknowledged
      IO_NewFault : Bool;   // Flag to start fault indicator (Lamp, Horn)
      IO_FaultAtStation : Bool;   // Fault at station active
      IO_PartShotNoNew : Int;
   END_VAR
   VAR_TEMP
      TempAmountTools : Word;
      TempStationNo : Int;
      Temp_EnableCycle : Bool;
      MH_No : Int;
      Temp_WK_No : Word;
      TempStationNoINT : Int;
      TmpActToolNo : Int;
      pDB : ANY;
      pAny AT pDB : Struct
         S7Code : Byte;
         DataType : Byte;
         Length : Int;
         DBNumber : Int;
         ByteAddressMSB : Word;
         ByteAddressLSB : Word;
      END_STRUCT;
      TmpMHatThisMachine : Bool;
      TmpDBNr : Int;
      TmpDBBAdress : Int;
      TmpBitAddress : Word;
      TmpS7Code : Byte;
      TmpDataType : Byte;
      MHNoShift : DWord;
      MHNoBinary : DWord;
      TmpDBBAdress_1 : Int;
      TmpDBBAdress_2 : Word;
      TmpToolNo : Int;
      TmpMachineNumber : Int;
   END_VAR
BEGIN
   //-----------------------------------------------------------------
   // Get values of tool and foaming data at foamingstation 
   // 19.02.13 HK
   //-----------------------------------------------------------------

   //-----------------------------------------------------------------
   //Set variabbles
   //-----------------------------------------------------------------
   #TmpMachineNumber := 1;//#IN_MachineNo ;
   #TmpMHatThisMachine := 0;
   #TmpActToolNo := 0;

   // Just for TEST please delete after testing
   // ------------------------------------------
   //  "DB009_Faults".Faults_Grp_1_at_PLC_M1 := FALSE;

   //------------------------------------------------------------------
   // Get station no. from FB110
   // -----------------------------------------------------------------
   #TempStationNo := WORD_TO_INT("DB110_Interf_Program_M1".Program_No_01);

   //-----------------------------------------------------------------
   // Acknowledge faults
   // ----------------------------------------------------------------
   IF #IN_ResetFaults  THEN
     #IO_Faults.FLT_NewNoTooEarly := False;
     #IO_Faults.FLT_WRongStationNumber := False; 
     #IO_Faults.FLT_WrongToolNumber := False;
     #IO_Faults.FLT_WrongMixingheadNumber := False;
     #IO_Faults.Reserve3 := False;
   END_IF;

   //------------------------------------------------------------------
   // Fault new station number too early
   // -----------------------------------------------------------------
   IF  #TempStationNo > 0                   AND
       ("DB619_State_MPart".Cycle[#TmpMachineNumber].PressurizeTimeRuns OR
       "DB619_State_MPart".Cycle[#TmpMachineNumber].CtrlChangeTimeRuns OR
       "DB619_State_MPart".Cycle[#TmpMachineNumber].running)           AND
       ("DB619_State_MPart".ToolMa[#TmpMachineNumber].StationNo <> INT_TO_BYTE(#TempStationNo)) AND
       "DB619_State_MPart".ToolMa[#TmpMachineNumber].StationActive AND NOT
       #IO_Faults.FLT_NewNoTooEarly  
   THEN 
         #IO_Faults.FLT_NewNoTooEarly := True;
         #IO_NewFault := True;
   END_IF;

   //------------------------------------------------------------------
   // Reset partshot no and flags
   // -----------------------------------------------------------------
   IF #TempStationNo = 0 AND 
       "DB619_State_MPart".ToolMa[#TmpMachineNumber].StationFinished OR NOT
       "DB619_State_MPart".Cycle[#TmpMachineNumber].Release
   THEN
       "DB619_State_MPart".ToolMa[#TmpMachineNumber].PartShot := 0;
       "DB619_State_MPart".ShotMa[#TmpMachineNumber].ShotData.MH_No := 0;
     #IO_PartShotNoNew:=  0;
     "DB619_State_MPart".ToolMa[#TmpMachineNumber].StationFinished:= False;
     "DB619_State_MPart".ToolMa[#TmpMachineNumber].StationActive := False;
     #TempStationNo := 0;
   END_IF;

   //---------------------------------------------------------------------
   // Get tool no., station no.; if station no. > 0 -> set Station active 
   // --------------------------------------------------------------------
   IF #TempStationNo > 0   AND
       #TempStationNo < "AmountAllocationAutomatic"  AND
     "DB619_State_MPart".ToolMa[#TmpMachineNumber].PartShot = 0 AND NOT
     #IO_Faults.FLT_WrongToolNumber                         AND NOT
     #IO_Faults.FLT_WrongMixingheadNumber                   AND NOT
     #IO_Faults.FLT_NewNoTooEarly  
   THEN
       IF ("DB110_Interf_Program_M1".Status_IF[1].IF_is_on_1_Position OR "DB110_Interf_Program_M1".Test_M01.Test_runs) AND "DB123_MH_IO_Signals".MH[1].IN.MH_Manual_Mode AND
           (#TempStationNo > 0 AND #TempStationNo < 101) THEN
           "DB619_State_MPart".ToolMa[#TmpMachineNumber].ToolNo := "DB941_Tool_alloc_manual_MH".MH[1].Alloc_stationTool[#TempStationNo];

       ELSIF "DB110_Interf_Program_M1".Status_IF[2].IF_is_on_1_Position AND "DB123_MH_IO_Signals".MH[2].IN.MH_Manual_Mode AND
           (#TempStationNo > 0 AND #TempStationNo < 101) THEN
           "DB619_State_MPart".ToolMa[#TmpMachineNumber].ToolNo := "DB941_Tool_alloc_manual_MH".MH[2].Alloc_stationTool[#TempStationNo];

       ELSIF "DB110_Interf_Program_M1".Status_IF[3].IF_is_on_1_Position AND "DB123_MH_IO_Signals".MH[3].IN.MH_Manual_Mode AND
           (#TempStationNo > 0 AND #TempStationNo < 101) THEN
           "DB619_State_MPart".ToolMa[#TmpMachineNumber].ToolNo := "DB941_Tool_alloc_manual_MH".MH[3].Alloc_stationTool[#TempStationNo];

       ELSIF "DB110_Interf_Program_M1".Status_IF[4].IF_is_on_1_Position AND "DB123_MH_IO_Signals".MH[4].IN.MH_Manual_Mode AND
           (#TempStationNo > 0 AND #TempStationNo < 101) THEN
           "DB619_State_MPart".ToolMa[#TmpMachineNumber].ToolNo := "DB941_Tool_alloc_manual_MH".MH[4].Alloc_stationTool[#TempStationNo];

       ELSIF "DB110_Interf_Program_M1".Status_IF[5].IF_is_on_1_Position AND "DB123_MH_IO_Signals".MH[5].IN.MH_Manual_Mode AND
           (#TempStationNo > 0 AND #TempStationNo < 101) THEN
           "DB619_State_MPart".ToolMa[#TmpMachineNumber].ToolNo := "DB941_Tool_alloc_manual_MH".MH[5].Alloc_stationTool[#TempStationNo];

       ELSIF "DB110_Interf_Program_M1".Status_IF[6].IF_is_on_1_Position AND "DB123_MH_IO_Signals".MH[6].IN.MH_Manual_Mode AND
           (#TempStationNo > 0 AND #TempStationNo < 101) THEN
           "DB619_State_MPart".ToolMa[#TmpMachineNumber].ToolNo := "DB941_Tool_alloc_manual_MH".MH[6].Alloc_stationTool[#TempStationNo];

       ELSIF "DB110_Interf_Program_M1".Status_IF[7].IF_is_on_1_Position AND "DB123_MH_IO_Signals".MH[7].IN.MH_Manual_Mode AND
           (#TempStationNo > 0 AND #TempStationNo < 101) THEN
           "DB619_State_MPart".ToolMa[#TmpMachineNumber].ToolNo := "DB941_Tool_alloc_manual_MH".MH[7].Alloc_stationTool[#TempStationNo];

       ELSIF "DB110_Interf_Program_M1".Status_IF[8].IF_is_on_1_Position AND "DB123_MH_IO_Signals".MH[8].IN.MH_Manual_Mode AND
           (#TempStationNo > 0 AND #TempStationNo < 101) THEN
           "DB619_State_MPart".ToolMa[#TmpMachineNumber].ToolNo := "DB941_Tool_alloc_manual_MH".MH[8].Alloc_stationTool[#TempStationNo];

       ELSIF "DB110_Interf_Program_M1".Status_IF[9].IF_is_on_1_Position AND "DB123_MH_IO_Signals".MH[9].IN.MH_Manual_Mode AND
           (#TempStationNo > 0 AND #TempStationNo < 101) THEN
           "DB619_State_MPart".ToolMa[#TmpMachineNumber].ToolNo := "DB941_Tool_alloc_manual_MH".MH[9].Alloc_stationTool[#TempStationNo];

       ELSIF "DB110_Interf_Program_M1".Status_IF[10].IF_is_on_1_Position AND "DB123_MH_IO_Signals".MH[10].IN.MH_Manual_Mode AND
           (#TempStationNo > 0 AND #TempStationNo < 101) THEN
           "DB619_State_MPart".ToolMa[#TmpMachineNumber].ToolNo := "DB941_Tool_alloc_manual_MH".MH[10].Alloc_stationTool[#TempStationNo];

       ELSIF "DB110_Interf_Program_M1".Status_IF[11].IF_is_on_1_Position AND "DB123_MH_IO_Signals".MH[11].IN.MH_Manual_Mode AND
           "DB123_MH_IO_Signals".MH[11].IN.MH_Start AND (#TempStationNo > 0 AND #TempStationNo < 101) THEN
           "DB619_State_MPart".ToolMa[#TmpMachineNumber].ToolNo := "DB941_Tool_alloc_manual_MH".MH[11].Alloc_stationTool[#TempStationNo];

       ELSIF "DB110_Interf_Program_M1".Status_IF[12].IF_is_on_1_Position AND "DB123_MH_IO_Signals".MH[12].IN.MH_Manual_Mode AND
           (#TempStationNo > 0 AND #TempStationNo < 101) THEN
           "DB619_State_MPart".ToolMa[#TmpMachineNumber].ToolNo := "DB941_Tool_alloc_manual_MH".MH[12].Alloc_stationTool[#TempStationNo];

       ELSIF "DB110_Interf_Program_M1".Status_IF[13].IF_is_on_1_Position AND "DB123_MH_IO_Signals".MH[13].IN.MH_Manual_Mode AND
           (#TempStationNo > 0 AND #TempStationNo < 101) THEN
           "DB619_State_MPart".ToolMa[#TmpMachineNumber].ToolNo := "DB941_Tool_alloc_manual_MH".MH[13].Alloc_stationTool[#TempStationNo];

       ELSIF "DB110_Interf_Program_M1".Status_IF[14].IF_is_on_1_Position AND "DB123_MH_IO_Signals".MH[14].IN.MH_Manual_Mode AND
           (#TempStationNo > 0 AND #TempStationNo < 101) THEN
           "DB619_State_MPart".ToolMa[#TmpMachineNumber].ToolNo := "DB941_Tool_alloc_manual_MH".MH[14].Alloc_stationTool[#TempStationNo];

       ELSIF "DB110_Interf_Program_M1".Status_IF[15].IF_is_on_1_Position AND "DB123_MH_IO_Signals".MH[15].IN.MH_Manual_Mode AND
           (#TempStationNo > 0 AND #TempStationNo < 101) THEN
           "DB619_State_MPart".ToolMa[#TmpMachineNumber].ToolNo := "DB941_Tool_alloc_manual_MH".MH[15].Alloc_stationTool[#TempStationNo];

